screen "7161_RecipeSetpoints_STRING" 1280x715, template "7xxx_Formats"
   Button "rec_BaseScreenLocked" at 0,0 size 1280x715; TextOff 'Text'
      Visibility <- "bo_System_BaseScreenLocked"
   ScreenModuleView "Setpoint_Display_String_2" at 4,166 size 1090x44; ScreenModuleType ""
      on Guid_{11997190-50501}: function_efd93a16("pop_recipes_STRING", 200, 50, -1, -1, 1); SetTag("CPG_Recipe_Management.popupTrackers[3]", 1)
      Guid_{11997190-47977} <- "CPG_Recipe_Management.setpointsArray_STRING[1]"
      Guid_{11997190-76362} <- "[1]"
   ScreenModuleView "Setpoint_Display_String_1" at 4,132 size 1090x44; ScreenModuleType ""
      on Guid_{11997190-50501}: function_efd93a16("pop_recipes_STRING", 200, 50, -1, -1, 1); SetTag("CPG_Recipe_Management.popupTrackers[3]", 0)
      Guid_{11997190-47977} <- "CPG_Recipe_Management.setpointsArray_STRING[0]"
      Guid_{11997190-76362} <- "[0]"
   ScreenModuleView "Setpoint_Display_String_3" at 4,200 size 1090x44; ScreenModuleType ""
      on Guid_{11997190-50501}: function_efd93a16("pop_recipes_STRING", 200, 50, -1, -1, 1); SetTag("CPG_Recipe_Management.popupTrackers[3]", 2)
      Guid_{11997190-47977} <- "CPG_Recipe_Management.setpointsArray_STRING[2]"
      Guid_{11997190-76362} <- "[2]"
   ScreenModuleView "Setpoint_Display_String_4" at 4,234 size 1090x44; ScreenModuleType ""
      on Guid_{11997190-50501}: function_efd93a16("pop_recipes_STRING", 200, 50, -1, -1, 1); SetTag("CPG_Recipe_Management.popupTrackers[3]", 3)
      Guid_{11997190-47977} <- "CPG_Recipe_Management.setpointsArray_STRING[3]"
      Guid_{11997190-76362} <- "[3]"
   ScreenModuleView "Setpoint_Display_String_5" at 4,268 size 1090x44; ScreenModuleType ""
      on Guid_{11997190-50501}: function_efd93a16("pop_recipes_STRING", 200, 50, -1, -1, 1); SetTag("CPG_Recipe_Management.popupTrackers[3]", 4)
      Guid_{11997190-47977} <- "CPG_Recipe_Management.setpointsArray_STRING[4]"
      Guid_{11997190-76362} <- "[4]"
   ScreenModuleView "Setpoint_Display_String_6" at 4,302 size 1090x44; ScreenModuleType ""
      on Guid_{11997190-50501}: function_efd93a16("pop_recipes_STRING", 200, 50, -1, -1, 1); SetTag("CPG_Recipe_Management.popupTrackers[3]", 5)
      Guid_{11997190-47977} <- "CPG_Recipe_Management.setpointsArray_STRING[5]"
      Guid_{11997190-76362} <- "[5]"
   ScreenModuleView "Setpoint_Display_String_7" at 4,336 size 1090x44; ScreenModuleType ""
      on Guid_{11997190-50501}: function_efd93a16("pop_recipes_STRING", 200, 50, -1, -1, 1); SetTag("CPG_Recipe_Management.popupTrackers[3]", 6)
      Guid_{11997190-47977} <- "CPG_Recipe_Management.setpointsArray_STRING[6]"
      Guid_{11997190-76362} <- "[6]"
   ScreenModuleView "Setpoint_Display_String_8" at 4,370 size 1090x44; ScreenModuleType ""
      on Guid_{11997190-50501}: function_efd93a16("pop_recipes_STRING", 200, 50, -1, -1, 1); SetTag("CPG_Recipe_Management.popupTrackers[3]", 7)
      Guid_{11997190-47977} <- "CPG_Recipe_Management.setpointsArray_STRING[7]"
      Guid_{11997190-76362} <- "[7]"
   ScreenModuleView "Setpoint_Display_String_9" at 4,404 size 1090x44; ScreenModuleType ""
      on Guid_{11997190-50501}: function_efd93a16("pop_recipes_STRING", 200, 50, -1, -1, 1); SetTag("CPG_Recipe_Management.popupTrackers[3]", 8)
      Guid_{11997190-47977} <- "CPG_Recipe_Management.setpointsArray_STRING[8]"
      Guid_{11997190-76362} <- "[8]"
   ScreenModuleView "Setpoint_Display_String_10" at 4,438 size 1090x44; ScreenModuleType ""
      on Guid_{11997190-50501}: function_efd93a16("pop_recipes_STRING", 200, 50, -1, -1, 1); SetTag("CPG_Recipe_Management.popupTrackers[3]", 9)
      Guid_{11997190-47977} <- "CPG_Recipe_Management.setpointsArray_STRING[9]"
      Guid_{11997190-76362} <- "[9]"
   ScreenModuleView "Setpoint_Display_String_11" at 4,472 size 1090x44; ScreenModuleType ""
      on Guid_{11997190-50501}: function_efd93a16("pop_recipes_STRING", 200, 50, -1, -1, 1); SetTag("CPG_Recipe_Management.popupTrackers[3]", 10)
      Guid_{11997190-47977} <- "CPG_Recipe_Management.setpointsArray_STRING[10]"
      Guid_{11997190-76362} <- "[10]"
   ScreenModuleView "Setpoint_Display_String_12" at 4,506 size 1090x44; ScreenModuleType ""
      on Guid_{11997190-50501}: function_efd93a16("pop_recipes_STRING", 200, 50, -1, -1, 1); SetTag("CPG_Recipe_Management.popupTrackers[3]", 11)
      Guid_{11997190-47977} <- "CPG_Recipe_Management.setpointsArray_STRING[11]"
      Guid_{11997190-76362} <- "[11]"
   TextField "Text field_9" at 125,40 size 227x25; Text 'RECIPE SETPOINTS - STRING / Rezeptur Sollwerte - STRING'
   Button "Button_3" at 160,555 size 78x45; TextOff 'Text'; PictureOff "Up_Arrow"
      on Release: function_b9b71300("CPG_Recipe_Management.currentPages[3]", 1)
   Button "Button_4" at 287,555 size 78x45; TextOff 'Text'; PictureOff "Down_Arrow"
      on Release: function_dd21b452("CPG_Recipe_Management.currentPages[3]", 1)
   TextField "Text field_10" at 35,565 size 126x25; Text 'Pg Up/Down / Seite vor/zurück'
   IOField "I/O field_3" at 446,565 size 35x25; FormatPattern 999
      ProcessValue <- "CPG_Recipe_Management.currentPages[3]"
   TextField "Text field_13" at 381,565 size 60x25; Text 'Page # / Seite #'
   TextField "Text field_14" at 488,565 size 32x25; Text 'of / von'
   IOField "I/O field_4" at 534,564 size 37x27; FormatPattern 999
      ProcessValue <- "CPG_Recipe_Management.maxPages[3]"
   TextField "Text field_2" at 35,93 size 115x25; Text 'Setpoint Name / Sollwert-Name'
   TextField "Text field_6" at 243,83 size 72x46; Text 'Current Value Aktueller Wert'
   TextField "Text field_7" at 384,93 size 32x25; Text 'Min'
   TextField "Text field_4" at 506,93 size 36x25; Text 'Max'
   IOField "I/O field_9" at 757,42 size 53x36; FormatPattern 999
      ProcessValue <- "RecipeID_A"
   IOField "I/O field_10" at 883,42 size 53x36; FormatPattern 999
      ProcessValue <- "RecipeID_B"
   IOField "I/O field_11" at 998,42 size 53x36; FormatPattern 999
      ProcessValue <- "RecipeID_C"
   IOField "I/O field_13" at 550,83 size 187x22; FormatPattern ????????????????????
      ProcessValue <- "CurrentRecipeName"
   IOField "I/O field_14" at 907,104 size 187x22; FormatPattern ????????????????????
      ProcessValue <- "RecipeName_C"
   IOField "I/O field_15" at 816,83 size 187x22; FormatPattern ????????????????????
      ProcessValue <- "RecipeName_B"
   IOField "I/O field_16" at 690,103 size 187x23; FormatPattern ????????????????????
      ProcessValue <- "RecipeName_A"
   TextField "Text field_1" at 748,15 size 98x25; Text 'Recipe A / Datensatz A'
   TextField "Text field_3" at 874,15 size 97x25; Text 'Recipe B / Datensatz B'
   TextField "Text field_8" at 989,15 size 97x25; Text 'Recipe C / Datensatz C'
   Group "Group" at 588,37 size 110x46
   TextField "Text field_5" at 588,37 size 88x46; Text 'Current Recipe: Aktueller Datensatz:'
   IOField "I/O field_12" at 663,48 size 35x25; FormatPattern 999
      ProcessValue <- "CurrentRecipeID"

screen "6001_SystemDiagnostic" 1280x715, template "6xxx_Diagnostics"
   SysDiagControl "ctrlSystemDiagnostics" at 15,15 size 1035x595
   Button "btnSystemDiagnosticsVerticalScrollUp" at 1050,70 size 40x30; TextOff 'Text'; PictureOff "icn-scroll-up-20x11"
      on Release: function_b22acb07("ctrlSystemDiagnostics")
   Button "btnSystemDiagnosticsVerticalScrollDown" at 1050,529 size 40x30; TextOff 'Text'; PictureOff "icn-scroll-down-20x11"
      on Release: function_b8b2ebe3("ctrlSystemDiagnostics")
   SysDiagControl "ctrlSystemDiagnosticsLocked" at 15,15 size 1035x595
      Visibility <- "bo_System_BaseScreenLocked"
   Rectangle "recBaseScreenLocked" at 0,0 size 1280x708
      Visibility <- "bo_System_BaseScreenLocked"

screen "6041_WebDiagnostic" 1280x715, template "6xxx_Diagnostics"
   HTMLBrowser "ctrlHTMLBrowser" at 16,16 size 1073x531
      Address <- "str_Diagnostic_WebURL"
   Button "btnWebServerPLC" at 15,560 size 125x50; TextOff 'PLC / SPS'
      on Release: SetTag("str_Diagnostic_WebURL", '192.168.0.1')
   Rectangle "recBaseScreenLocked" at 0,0 size 1280x708
      Visibility <- "bo_System_BaseScreenLocked"

Template "1xxx_MachineControl" 1280x715
   ScreenModuleView "fcpBodyBar" at 5,5 size 1270x615; Guid_{11997190-53329} 'Up & Downstream'; Guid_{11997190-53335} 'OMAC Times OMAC Zeiten Timers / OEE'; Guid_{11997190-53325} 'Overview / Übersicht / Equipment view'; Guid_{11997190-53331} 'OMAC State Model OMAC Statusmodell OMAC State Model'; Guid_{11997190-53337} 'OEE / Manual CMD's'; Guid_{11997190-53333} 'OMAC PackTags PackTags'; Guid_{11997190-53339} 'Manual Commands Manuelle Kommandos PDI Interface'; ScreenModuleType ""
      on Guid_{11997190-53582}: ActivateScreen("1201_OEE", 0)
      on Guid_{11997190-53576}: ActivateScreen("1081_OMACStateModel", 0)
      on Guid_{11997190-53580}: ActivateScreen("1161_OMACTimes", 0)
      on Guid_{11997190-53584}: ActivateScreen("1241_ManualCommands", 0)
      on Guid_{11997190-53578}: ActivateScreen("1121_OMACPackTags", 0)
      on Guid_{11997190-53574}: ActivateScreen("1041_Up&Downstream", 0)
      on Guid_{11997190-53572}: ActivateScreen("1001_EquipmentView1", 0)
      Guid_{11997190-62386} <- "HMI_Data.HMICurrentScreenID"
      Guid_{11997190-53044} <- "i16_1000_MachineControl_SecondNavMaxTopics"
   ScreenModuleView "fcpBottomBar" at 5,625 size 1270x85; ScreenModuleType ""
      on Guid_{11997190-126458}: function_efd93a16("pop_UserLogin", 437, 285, 1, -1, 1)
      on Guid_{11997190-96858}: ActivateScreen("6001_SystemDiagnostic", 0)
      on Guid_{11997190-96860}: ActivateScreen("7001_RecipeControl", 0)
      on Guid_{11997190-126452}: "sub_OpenPrevScreen"()
      on Guid_{11997190-96848}: ActivateScreen("1001_EquipmentView1", 0)
      on Guid_{11997190-96850}: ActivateScreen("2001_Settings", 0)
      on Guid_{11997190-96852}: ActivateScreen("3001_AlarmOverview", 0)
      Guid_{11997190-60598} <- "HMI_Data.HMICurrentScreenID"
   Button "btnCntrlCmdStart" at 835,638 size 70x70; TextOff 'Text'; PictureOff "icn-omac-start"
      on Release: ResetBit("HMI_Data.CMDs.PB_Start")
      on Press: SetBit("HMI_Data.CMDs.PB_Start")
      Appearance <- "HMI_Data.CMDs.PB_Start"
   Button "btnCntrlCmdStop" at 910,638 size 70x70; TextOff 'Text'; PictureOff "icn-omac-stop"
      on Release: ResetBit("HMI_Data.CMDs.PB_Stop")
      on Press: SetBit("HMI_Data.CMDs.PB_Stop")
      Appearance <- "HMI_Data.CMDs.PB_Stop"
   Button "btnCntrlCmdReset" at 985,638 size 70x70; TextOff 'Text'; PictureOff "icn-omac-reset"
      on Release: ResetBit("HMI_Data.CMDs.PB_Reset")
      on Press: SetBit("HMI_Data.CMDs.PB_Reset")
      Appearance <- "HMI_Data.CMDs.PB_Reset"
   Switch "Switch_EStop" at 1126,517 size 132x58; CaptionText 'Switch'; TextOff 'E-Stop Released Not-Halt Quittiert'; TextOn 'E-Stop Pressed Not-Halt Aktiv'
      ProcessValue <- "HMI_Data_CPG.CMDs.PB_EStop"
      Appearance <- "HMI_Data_CPG.CMDs.PB_EStop"

Template "2xxx_Settings" 1280x715
   ScreenModuleView "fcpBodyBar" at 5,5 size 1270x615; Guid_{11997190-53325} 'Station A / Estacion A'; Guid_{11997190-53331} 'Benutzer- verwaltung'; Guid_{11997190-53329} 'System Functions System- funktionen Estacion B'; ScreenModuleType ""
      on Guid_{11997190-53576}: ActivateScreen("2081_UserManagement", 0)
      on Guid_{11997190-53574}: ActivateScreen("2041_SystemFunctions", 0)
      on Guid_{11997190-53572}: ActivateScreen("2001_Settings", 0)
      Guid_{11997190-62386} <- "HMI_Data.HMICurrentScreenID"
      Guid_{11997190-53044} <- "i16_2000_Settings_SecondNavMaxTopics"
   ScreenModuleView "fcpBottomBar" at 5,625 size 1270x85; ScreenModuleType ""
      on Guid_{11997190-126458}: function_efd93a16("pop_UserLogin", 437, 285, 1, -1, 1)
      on Guid_{11997190-96858}: ActivateScreen("6001_SystemDiagnostic", 0)
      on Guid_{11997190-96860}: ActivateScreen("7001_RecipeControl", 0)
      on Guid_{11997190-126452}: "sub_OpenPrevScreen"()
      on Guid_{11997190-96848}: ActivateScreen("1001_EquipmentView1", 0)
      on Guid_{11997190-96850}: ActivateScreen("2001_Settings", 0)
      on Guid_{11997190-96852}: ActivateScreen("3001_AlarmOverview", 0)
      Guid_{11997190-60598} <- "HMI_Data.HMICurrentScreenID"
   Button "btnCntrlCmdStart" at 835,638 size 70x70; TextOff 'Text'; PictureOff "icn-omac-start"
      on Release: ResetBit("HMI_Data.CMDs.PB_Start")
      on Press: SetBit("HMI_Data.CMDs.PB_Start")
      Appearance <- "HMI_Data.CMDs.PB_Start"
   Button "btnCntrlCmdStop" at 910,638 size 70x70; TextOff 'Text'; PictureOff "icn-omac-stop"
      on Release: ResetBit("HMI_Data.CMDs.PB_Stop")
      on Press: SetBit("HMI_Data.CMDs.PB_Stop")
      Appearance <- "HMI_Data.CMDs.PB_Stop"
   Button "btnCntrlCmdReset" at 985,638 size 70x70; TextOff 'Text'; PictureOff "icn-omac-reset"
      on Release: ResetBit("HMI_Data.CMDs.PB_Reset")
      on Press: SetBit("HMI_Data.CMDs.PB_Reset")
      Appearance <- "HMI_Data.CMDs.PB_Reset"

Template "3xxx_Alarms&Events" 1280x715
   ScreenModuleView "fcpBodyBar" at 5,5 size 1270x615; Guid_{11997190-53329} 'Alarm Events / Alarmmeldungen'; Guid_{11997190-53335} 'Pareto Alarm Tracking'; Guid_{11997190-53325} 'Event Overview / Meldeübersicht'; Guid_{11997190-53331} 'Warning Events / Warnmeldungen / Eventos de advertencia'; Guid_{11997190-53333} 'HMI Events / HMI Meldungen'; ScreenModuleType ""
      on Guid_{11997190-53576}: ActivateScreen("3081_WarningEvents", 0)
      on Guid_{11997190-53574}: ActivateScreen("3041_AlarmEvents", 0)
      on Guid_{11997190-53578}: ActivateScreen("3121_HMI_Alarms", 0)
      on Guid_{11997190-53580}: ActivateScreen("3161_ParetoAlarmData", 0)
      on Guid_{11997190-53572}: ActivateScreen("3001_AlarmOverview", 0)
      Guid_{11997190-62386} <- "HMI_Data.HMICurrentScreenID"
      Guid_{11997190-53044} <- "i16_3000_Alarms&Events_SecondNavMaxTopics"
   ScreenModuleView "fcpBottomBar" at 5,625 size 1270x85; ScreenModuleType ""
      on Guid_{11997190-126458}: function_efd93a16("pop_UserLogin", 437, 285, 1, -1, 1)
      on Guid_{11997190-96858}: ActivateScreen("6001_SystemDiagnostic", 0)
      on Guid_{11997190-96860}: ActivateScreen("7001_RecipeControl", 0)
      on Guid_{11997190-126452}: "sub_OpenPrevScreen"()
      on Guid_{11997190-96848}: ActivateScreen("1001_EquipmentView1", 0)
      on Guid_{11997190-96850}: ActivateScreen("2001_Settings", 0)
      on Guid_{11997190-96852}: ActivateScreen("3001_AlarmOverview", 0)
      Guid_{11997190-60598} <- "HMI_Data.HMICurrentScreenID"
   Button "btnCntrlCmdStart" at 835,638 size 70x70; TextOff 'Text'; PictureOff "icn-omac-start"
      on Release: ResetBit("HMI_Data.CMDs.PB_Start")
      on Press: SetBit("HMI_Data.CMDs.PB_Start")
      Appearance <- "HMI_Data.CMDs.PB_Start"
   Button "btnCntrlCmdStop" at 910,638 size 70x70; TextOff 'Text'; PictureOff "icn-omac-stop"
      on Release: ResetBit("HMI_Data.CMDs.PB_Stop")
      on Press: SetBit("HMI_Data.CMDs.PB_Stop")
      Appearance <- "HMI_Data.CMDs.PB_Stop"
   Button "btnCntrlCmdReset" at 985,638 size 70x70; TextOff 'Text'; PictureOff "icn-omac-reset"
      on Release: ResetBit("HMI_Data.CMDs.PB_Reset")
      on Press: SetBit("HMI_Data.CMDs.PB_Reset")
      Appearance <- "HMI_Data.CMDs.PB_Reset"

Template "6xxx_Diagnostics" 1280x715
   ScreenModuleView "fcpBodyBar" at 5,5 size 1270x615; Guid_{11997190-53325} 'System Diagnostic System- diagnose Diagnóstico del sistema'; Guid_{11997190-53329} 'Web Diagnostic Web- diagnose Diagnóstico web'; ScreenModuleType ""
      on Guid_{11997190-53574}: ActivateScreen("6041_WebDiagnostic", 0)
      on Guid_{11997190-53572}: ActivateScreen("6001_SystemDiagnostic", 0)
      Guid_{11997190-62386} <- "HMI_Data.HMICurrentScreenID"
      Guid_{11997190-53044} <- "i16_6000_Diagnostics_SecondNavMaxTopics"
   ScreenModuleView "fcpBottomBar" at 5,625 size 1270x85; ScreenModuleType ""
      on Guid_{11997190-126458}: function_efd93a16("pop_UserLogin", 437, 285, 1, -1, 1)
      on Guid_{11997190-96858}: ActivateScreen("6001_SystemDiagnostic", 0)
      on Guid_{11997190-96860}: ActivateScreen("7001_RecipeControl", 0)
      on Guid_{11997190-126452}: "sub_OpenPrevScreen"()
      on Guid_{11997190-96848}: ActivateScreen("1001_EquipmentView1", 0)
      on Guid_{11997190-96850}: ActivateScreen("2001_Settings", 0)
      on Guid_{11997190-96852}: ActivateScreen("3001_AlarmOverview", 0)
      Guid_{11997190-60598} <- "HMI_Data.HMICurrentScreenID"
   Button "btnCntrlCmdStart" at 835,638 size 70x70; TextOff 'Text'; PictureOff "icn-omac-start"
      on Release: ResetBit("HMI_Data.CMDs.PB_Start")
      on Press: SetBit("HMI_Data.CMDs.PB_Start")
      Appearance <- "HMI_Data.CMDs.PB_Start"
   Button "btnCntrlCmdStop" at 910,638 size 70x70; TextOff 'Text'; PictureOff "icn-omac-stop"
      on Release: ResetBit("HMI_Data.CMDs.PB_Stop")
      on Press: SetBit("HMI_Data.CMDs.PB_Stop")
      Appearance <- "HMI_Data.CMDs.PB_Stop"
   Button "btnCntrlCmdReset" at 985,638 size 70x70; TextOff 'Text'; PictureOff "icn-omac-reset"
      on Release: ResetBit("HMI_Data.CMDs.PB_Reset")
      on Press: SetBit("HMI_Data.CMDs.PB_Reset")
      Appearance <- "HMI_Data.CMDs.PB_Reset"

Template "7xxx_Formats" 1280x715
   ScreenModuleView "fcpBodyBar" at 5,5 size 1270x615; Guid_{11997190-53329} 'REAL Sollwerte'; Guid_{11997190-53335} 'STRING Sollwerte'; Guid_{11997190-53325} 'Recipe Control Rezepturverwaltung'; Guid_{11997190-53331} 'DINT Sollwerte'; Guid_{11997190-53333} 'BOOL Sollwerte'; ScreenModuleType ""
      on Guid_{11997190-53576}: ActivateScreen("7081_RecipeSetpoints_DINT", 0)
      on Guid_{11997190-53580}: ActivateScreen("7161_RecipeSetpoints_STRING", 0)
      on Guid_{11997190-53578}: ActivateScreen("7121_RecipeSetpoints_BOOL", 0)
      on Guid_{11997190-53574}: ActivateScreen("7041_RecipeSetpoints_REAL", 0)
      on Guid_{11997190-53572}: ActivateScreen("7001_RecipeControl", 0)
      Guid_{11997190-62386} <- "HMI_Data.HMICurrentScreenID"
      Guid_{11997190-53044} <- "i16_7000_Formats_SecondNavMaxTopics"
   ScreenModuleView "fcpBottomBar" at 5,625 size 1270x85; ScreenModuleType ""
      on Guid_{11997190-126458}: function_efd93a16("pop_UserLogin", 437, 285, 1, -1, 1)
      on Guid_{11997190-96858}: ActivateScreen("6001_SystemDiagnostic", 0)
      on Guid_{11997190-96860}: ActivateScreen("7001_RecipeControl", 0)
      on Guid_{11997190-126452}: "sub_OpenPrevScreen"()
      on Guid_{11997190-96848}: ActivateScreen("1001_EquipmentView1", 0)
      on Guid_{11997190-96850}: ActivateScreen("2001_Settings", 0)
      on Guid_{11997190-96852}: ActivateScreen("3001_AlarmOverview", 0)
      Guid_{11997190-60598} <- "HMI_Data.HMICurrentScreenID"
   Button "btnCntrlCmdStart" at 835,638 size 70x70; TextOff 'Text'; PictureOff "icn-omac-start"
      on Release: ResetBit("HMI_Data.CMDs.PB_Start")
      on Press: SetBit("HMI_Data.CMDs.PB_Start")
      Appearance <- "HMI_Data.CMDs.PB_Start"
   Button "btnCntrlCmdStop" at 910,638 size 70x70; TextOff 'Text'; PictureOff "icn-omac-stop"
      on Release: ResetBit("HMI_Data.CMDs.PB_Stop")
      on Press: SetBit("HMI_Data.CMDs.PB_Stop")
      Appearance <- "HMI_Data.CMDs.PB_Stop"
   Button "btnCntrlCmdReset" at 985,638 size 70x70; TextOff 'Text'; PictureOff "icn-omac-reset"
      on Release: ResetBit("HMI_Data.CMDs.PB_Reset")
      on Press: SetBit("HMI_Data.CMDs.PB_Reset")
      Appearance <- "HMI_Data.CMDs.PB_Reset"

PopupScreen "pop_ErrorScreenNo" 405x230
   on GenerateScreen: SetBit("bo_System_BaseScreenLocked")
   on ClearScreen: ResetBit("bo_System_BaseScreenLocked")
   Button "btnClose" at 140,170 size 125x50; TextOff 'Close / Schließen'
      on Click: function_efd93a16("pop_ErrorScreenNo", 0, 0, 0, -1, 1)
   TextField "txtMessage" at 10,65 size 390x105; Text 'The screen number could not be determined! Please check the screen name. Die Bildnummer konnte nicht ermittelt werden! Bitte überprüfen Sie den Bildnamen. The Screen name has the wrong Style'
   Button "btnHeader" at 3,3 size 399x60; TextOff 'System Error / Systemfehler'

PopupScreen "pop_UserLogin" 405x230
   on GenerateScreen: SetBit("bo_System_BaseScreenLocked")
   on ClearScreen: ResetBit("bo_System_BaseScreenLocked")
   Button "btnLogOff" at 10,170 size 125x50; TextOff 'Log off / Ausloggen / Desconectarse'
      on Release: function_efd93a16("pop_UserLogin", 0, 0, 0, -1, 1); function_f23ef4c9()
   Button "btnChangeUser" at 140,170 size 125x50; TextOff 'Change User Benutzer- wechsel'
      on Release: function_efd93a16("pop_UserLogin", 0, 0, 0, -1, 1); function_a2a04561()
   Button "btnClose" at 270,170 size 125x50; TextOff 'Close / Schließen'
      on Release: function_efd93a16("pop_UserLogin", 0, 0, 0, -1, 1)
   TextField "txtMessage" at 10,65 size 390x105; Text 'Log off or change user? / Ausloggen oder Benutzerwechsel?'
   Button "btnHeader" at 3,3 size 399x60; TextOff 'User Management / Benutzerverwaltung'

PopupScreen "pop_recipes_BOOL" 645x584
   ScreenModuleView "Bool Popup_1_1" at 2,1 size 640x579; ScreenModuleType ""
      on Guid_{11997190-50035}: ActivateScreen("7121_RecipeSetpoints_BOOL", 0)
      Guid_{11997190-48328} <- "CPG_Recipe_Management.setpointPopup_BOOL"
      Guid_{11997190-42630} <- "CPG_RecipeCfg.recipeControl"

PopupScreen "pop_recipes_DINT" 645x584
   ScreenModuleView "Dint Popup_1" at 0,0 size 640x579; ScreenModuleType ""
      on Guid_{11997190-50035}: ActivateScreen("7081_RecipeSetpoints_DINT", 0)
      Guid_{11997190-48328} <- "CPG_Recipe_Management.setpointPopup_DINT"
      Guid_{11997190-42630} <- "CPG_RecipeCfg.recipeControl"

PopupScreen "pop_recipes_REAL" 642x581
   ScreenModuleView "Real Popup_1" at 0,0 size 640x579; ScreenModuleType ""
      on Guid_{11997190-50035}: ActivateScreen("7041_RecipeSetpoints_REAL", 0)
      Guid_{11997190-48328} <- "CPG_Recipe_Management.setpointPopup_REAL"
      Guid_{11997190-42630} <- "CPG_RecipeCfg.recipeControl"

PopupScreen "pop_recipes_STRING" 645x584
   ScreenModuleView "Popup_String_1" at 2,0 size 640x579; ScreenModuleType ""
      on Guid_{11997190-50035}: ActivateScreen("7161_RecipeSetpoints_STRING", 0)
      Guid_{11997190-48328} <- "CPG_Recipe_Management.setpointPopup_STRING"
      Guid_{11997190-42630} <- "CPG_RecipeCfg.recipeControl"

VB script "sub_SetScreenBrightness"
   '****************************************************************************************************************************
   '----------------------------------------------------------------------------------------------------------------------------
   ' Functionality : Changing the screen brightness with a defined increment size
   ' Run           : After a user change via the task scheduler
   ' Run system    : WinCC Comfort/Advanced Runtime V13
   '----------------------------------------------------------------------------------------------------------------------------
   ' Script parameters:
   '  Parameter        | Data type    | Description
   '  i16Offset        | INTEGER      | Specifies the increment by which the screen brightness is changed
   '----------------------------------------------------------------------------------------------------------------------------
   ' Change table:
   '  Version    | Date     | Creator         | Description
   '  01.00.00   | 18/06/18 | Briese, Mike    | Creation
   '----------------------------------------------------------------------------------------------------------------------------
   '****************************************************************************************************************************
   
   'Declaration
   Dim i16NewDisplayBrightness
   
   
   'Determine new value for screen brightness
   i16NewDisplayBrightness = SmartTags("i16_Settings_CurDisplayBrightness") + i16Offset
   
   'Check whether new value is within the limits
   '=> If No, then set to the corresponding limit value
   If i16NewDisplayBrightness < 20 Then
   	i16NewDisplayBrightness = 20
   ElseIf i16NewDisplayBrightness > 100 Then
   	i16NewDisplayBrightness = 100
   End If
   
   'Take over new value
   SmartTags("i16_Settings_CurDisplayBrightness") = i16NewDisplayBrightness
   e4c2bb66-d114-4215-9f74-4e7e992fb119 i16NewDisplayBrightness

VB script "sub_ScreenChanged"
   '****************************************************************************************************************************
   '----------------------------------------------------------------------------------------------------------------------------
   ' Functionality : Determining the screen number from the screen name
   ' Run           : After a screen change via the task scheduler
   ' Run system    : WinCC Comfort/Advanced Runtime V13
   '----------------------------------------------------------------------------------------------------------------------------
   ' Script parameters:
   '  Parameter        | Data type    | Description
   '                   |              |
   '----------------------------------------------------------------------------------------------------------------------------
   ' Change table:
   '  Version    | Date     | Creator         | Description
   '  01.00.00   | 18/06/18 | Briese, Mike    | Creation
   '----------------------------------------------------------------------------------------------------------------------------
   '****************************************************************************************************************************
   
   'Declaration
   Dim strCurScreenName, i16NewScreenID, i16Index
   
   
   'Determine screen number from screen name
   strCurScreenName = HmiRuntime.BaseScreenName
   i16NewScreenID = Mid(strCurScreenName, 1, 4)
   
   'Plausibility check of the determined screen number
   '=> if it is not plausible, show an error message and exit sub
   If Not IsNumeric(i16NewScreenID) Then
   	efd93a16-2665-4b85-bcb9-25eddcb7b6f4 pop_ErrorScreenNo, 437, 285, $3$hmiOn$, $3$hmiAnimationOff$, $3$hmiMedium$
   	SmartTags("HMI_Data.HMICurrentScreenID") = -1
   	Exit Sub
   End If 
   
   'Take over determined screen number
   SmartTags("HMI_Data.HMICurrentScreenID") = i16NewScreenID
   
   'Take over determined screen number to screen buffer for return function, if this is not active
   i16Index = SmartTags("i16_System_PrevScreenPointer")
   If SmartTags("bo_System_PrevScreenActive") Then
   	SmartTags("bo_System_PrevScreenActive") = False
   Else
   	If i16Index < UBound(SmartTags("arr_System_PrevScreenStorage")) Then
   		i16Index = i16Index + 1
   	Else
   		i16Index = 0
   	End If
   	SmartTags("i16_System_PrevScreenPointer") = i16Index
   	SmartTags("arr_System_PrevScreenStorage")(i16Index) = i16NewScreenID
   End If

VB script "sub_RuntimeStart"
   '****************************************************************************************************************************
   '----------------------------------------------------------------------------------------------------------------------------
   ' Functionality : This script contains all one-time actions that are to be executed after the runtime start
   ' Run           : Runtime start of HMI project
   ' Run system    : WinCC Comfort/Advanced Runtime V13
   '----------------------------------------------------------------------------------------------------------------------------
   ' Script parameters:
   '  Parameter        | Data type    | Description
   '                   |              |
   '----------------------------------------------------------------------------------------------------------------------------
   ' Change table:
   '  Version    | Date     | Creator         | Description
   '  01.00.00   | 18/06/18 | Briese, Mike    | Creation
   '----------------------------------------------------------------------------------------------------------------------------
   '****************************************************************************************************************************
   
   
   'Determine current user info
   sub_UserChanged
   
   'Open overview screen
   bec8f1e5-2ab1-45f6-ad91-1d37c469eb91 1001_EquipmentView1, 0

VB script "sub_OpenPrevScreen"
   '****************************************************************************************************************************
   '----------------------------------------------------------------------------------------------------------------------------
   ' Functionality : Open previous screen
   '                 An screen buffer is required for this function. 
   ' Run           : On demand
   ' Run system    : WinCC Comfort/Advanced Runtime V13
   '----------------------------------------------------------------------------------------------------------------------------
   ' Script parameters:
   '  Parameter        | Data type    | Description
   '                   |              |
   '----------------------------------------------------------------------------------------------------------------------------
   ' Change table:
   '  Version    | Date     | Creator         | Description
   '  01.00.00   | 18/06/18 | Briese, Mike    | Creation
   '----------------------------------------------------------------------------------------------------------------------------
   '****************************************************************************************************************************
   
   'Declaration
   Const strFctName = "sub_OpenPrevScreen"
   Dim i16CurBufferIndex, i16NewBufferIndex, i16ScreenID
   
   
   'Load number of previous screen from screen buffer
   i16CurBufferIndex = SmartTags("i16_System_PrevScreenPointer")
   If i16CurBufferIndex > 0 Then
   	i16NewBufferIndex = i16CurBufferIndex - 1
   Else
   	i16NewBufferIndex = UBound(SmartTags("arr_System_PrevScreenStorage"))
   End If
   
   'Check if screen buffer element contains a valid number
   '=> if no, then the function is terminated
   i16ScreenID = SmartTags("arr_System_PrevScreenStorage")(i16NewBufferIndex)
   If i16ScreenID = 0 Then Exit Sub
   
   'Reset current screen buffer element and accept new pointer
   SmartTags("arr_System_PrevScreenStorage")(i16CurBufferIndex) = 0
   SmartTags("i16_System_PrevScreenPointer") = i16NewBufferIndex
   
   'Set auxiliary flag for screen change function
   SmartTags("bo_System_PrevScreenActive") = True
   
   'Open previous screen
   acd163fa-ee86-4170-88da-c8d9ec58660c i16ScreenID, 0

VB script "sub_UserChanged"
   '****************************************************************************************************************************
   '----------------------------------------------------------------------------------------------------------------------------
   ' Functionality : Determining the screen number from the screen name
   '                 The associated group number/name and authorizations are determined according to the current user selection.
   '                 Afterwards, a '0' is entered at the current pointer position in the screen storage for the return function,
   '                 so that the new user cannot jump to the last called screens of the previous user. Finally, the overview
   '                 screen is opened.
   ' Run           : After a user change via the task scheduler
   ' Run system    : WinCC Comfort/Advanced Runtime V13
   '----------------------------------------------------------------------------------------------------------------------------
   ' Script parameters:
   '  Parameter        | Data type    | Description
   '                   |              |
   '----------------------------------------------------------------------------------------------------------------------------
   ' Change table:
   '  Version    | Date     | Creator         | Description
   '  01.00.00   | 18/06/18 | Briese, Mike    | Creation
   '----------------------------------------------------------------------------------------------------------------------------
   '****************************************************************************************************************************
   
   'Declaration
   Dim arrUserName, strUserName(2), strUserNamePart1, strUserNamePart2, strLoginData
   Dim i16Index
   
   'Determine current user name
   f41c6f6c-971d-4734-9362-16d81ac70597 str_System_CurUser
   If SmartTags("str_System_CurUser") = "" Then
   	SmartTags("str_System_CurUser") = "-"
   End If
   
   'Initialize current pointer index of the screen buffer for return function
   '=> to restart from here after changing users
   i16Index = SmartTags("i16_System_PrevScreenPointer")
   SmartTags("arr_System_PrevScreenStorage")(i16Index) = 0
   
   'Reset basic screen lock
   '=> required if incorrect login data has been entered
   SmartTags("bo_System_BaseScreenLocked") = False
   
   'Open overview screen
   bec8f1e5-2ab1-45f6-ad91-1d37c469eb91 1001_EquipmentView1, 0

scheduled task "ScreenChanged"
   on Action: "sub_ScreenChanged"()

scheduled task "UserChanged"
   on Action: "sub_UserChanged"()
*)

(* ===== HMI "HMI_RT_1" =====
system functions are stored by id; their names below are inferred from use

HMI tags "Default tag table"
   "testtag" : WString[10], internal

ScreenModuleEditorView "Popup_Real" 700x600
   Rectangle "Rectangle_2" at 113,186 size 434x39
      Visibility <- "Setpoint.SetpointChangeDisabled"
   TextField "NotAllowed Warning" at 131,194 size 398x23; Text 'Setpoint Changes Not Allowed in Current Machine State / Änderung im aktuellen Maschinenzustand nicht möglich'
      Visibility <- "Setpoint.SetpointChangeDisabled"
   Rectangle "Yellow" at 113,72 size 434x39
      Visibility <- "Setpoint.RecipeSetpointDiff"
   TextField "DetectDiff Warning" at 141,80 size 402x23; Text 'Current Setpoint Does Not Match Saved Recipe Value / Der aktuelle Sollwert entspricht nicht dem gespeicherten'
      Visibility <- "Setpoint.RecipeSetpointDiff"
   IOField "Current Num" at 69,346 size 46x26; FormatPattern 999
      ProcessValue <- "Control.CurrentRecipeID"
   IOField "NumA" at 69,388 size 46x26; FormatPattern 999
      ProcessValue <- "Control.RecipeID_A"
   IOField "NumB" at 69,429 size 46x26; FormatPattern 999
      ProcessValue <- "Control.RecipeID_B"
   IOField "NumC" at 69,471 size 46x26; FormatPattern 999
      ProcessValue <- "Control.RecipeID_C"
   TextField "Text field_5" at 239,305 size 112x23; Text 'Recipe Name / Datensatzname'
   TextField "Text field_6" at 517,305 size 44x23; Text 'Value / Wert'
   TextField "Text field_7" at 266,264 size 129x28; Text 'Recipe Values / Rezepturwert'
   IOField "CurrentValue_true" at 486,348 size 106x23; FormatPattern 9999999.999
      ProcessValue <- "Setpoint.CurrentRecipeValue"
   IOField "ValueA" at 486,390 size 106x25; FormatPattern 9999999.999
      ProcessValue <- "Setpoint.RecipeValueA"
   IOField "ValueB" at 486,431 size 106x23; FormatPattern 9999999.999
      ProcessValue <- "Setpoint.RecipeValueB"
   IOField "ValueC" at 486,473 size 106x23; FormatPattern 9999999.999
      ProcessValue <- "Setpoint.RecipeValueC"
   IOField "CurrentName" at 158,346 size 282x26; FormatPattern ??????????????????????????????
      ProcessValue <- "Control.CurrentRecipeName"
   IOField "NameA" at 158,388 size 282x26; FormatPattern ??????????????????????????????
      ProcessValue <- "Control.RecipeName_A"
   IOField "NameB" at 158,429 size 282x26; FormatPattern ??????????????????????????????
      ProcessValue <- "Control.RecipeName_B"
   IOField "NameC" at 158,471 size 282x26; FormatPattern ??????????????????????????????
      ProcessValue <- "Control.RecipeName_C"
   Group "Group" at 113,186 size 434x39
   Group "Group_1" at 113,72 size 434x39
   IOField "Setpoint Name" at 145,27 size 370x41; FormatPattern ????????????????????????????????
      ProcessValue <- "Setpoint.CurrentName"
   Button "Save Setpoint" at 429,233 size 154x60; TextOff 'Save Setpoint Value Sollwert Speichern'
      on Press: function_b14e0dd5("Setpoint.SaveSetpoint", 0)
   Button "Revert Setpoint" at 69,233 size 154x60; TextOff 'Revert Setpoint Value Sollwert Rücksetzen'
      on Press: function_b14e0dd5("Setpoint.RevertSetpoint", 0)
   Button "Close Button" at 79,519 size 502x60; TextOff 'CLOSE / Schließen'
   IOField "CurrentValue_true_1" at 206,153 size 132x26; FormatPattern 9999999.999
      ProcessValue <- "Setpoint.IN"
   TextField "Text field_1" at 79,307 size 36x23; Text '#'
   IOField "Max Value" at 464,154 size 106x23; FormatPattern 9999999.999
      ProcessValue <- "Setpoint.maxLimit"
   IOField "Min Value" at 93,154 size 106x23; FormatPattern 9999999.999
      ProcessValue <- "Setpoint.minLimit"
   Rectangle "Min Warning" at 94,147 size 104x36
      Visibility <- "Setpoint.minLimitReached"
   Rectangle "Max Warning" at 465,147 size 104x36
      Visibility <- "Setpoint.maxLimitReached"
   TextField "Text field_2" at 267,116 size 133x28; Text 'Current Value / Aktueller Wert'
   TextField "Text field_3" at 123,116 size 45x28; Text 'Min'
   TextField "Text field_4" at 494,116 size 45x28; Text 'Max'
   Group "Group_2" at 32,230 size 597x289
   Group "Group_3" at 345,153 size 112x23
   Rectangle "Rectangle_3" at 32,230 size 597x289
      Visibility <- "Setpoint.DisableRecipeControl"
   TextField "Text field_8" at 246,348 size 223x23; Text 'Recipe Control Disabled / Rezepturverwaltung deaktiviert'
      Visibility <- "Setpoint.DisableRecipeControl"
   TextField "Text field_10" at 345,153 size 112x23; Text '[ ]'
   IOField "Unit" at 353,153 size 96x23; FormatPattern ??????????
      ProcessValue <- "Setpoint.unit"
*)

(* ===== HMI "HMI_RT_1" =====
system functions are stored by id; their names below are inferred from use

HMI tags "Default tag table"
   "testtag" : WString[10], internal

ScreenModuleEditorView "Popup_String" 700x600
   Rectangle "Rectangle_2" at 113,154 size 434x39
      Visibility <- "Setpoint.SetpointChangeDisabled"
   TextField "NotAllowed Warning" at 131,162 size 398x23; Text 'Setpoint Changes Not Allowed in Current Machine State / Änderung im aktuellen Maschinenzustand nicht möglich'
      Visibility <- "Setpoint.SetpointChangeDisabled"
   Rectangle "Yellow" at 113,72 size 434x39
      Visibility <- "Setpoint.RecipeSetpointDiff"
   TextField "DetectDiff Warning" at 141,80 size 379x23; Text 'Current Setpoint Does Not Match Saved Recipe Value / Der aktuelle Sollwert entspricht dem gespeicherten'
      Visibility <- "Setpoint.RecipeSetpointDiff"
   IOField "Current Num" at 69,346 size 46x26; FormatPattern 999
      ProcessValue <- "Control.CurrentRecipeID"
   IOField "NumA" at 69,388 size 46x26; FormatPattern 999
      ProcessValue <- "Control.RecipeID_A"
   IOField "NumB" at 69,429 size 46x26; FormatPattern 999
      ProcessValue <- "Control.RecipeID_B"
   IOField "NumC" at 69,471 size 46x26; FormatPattern 999
      ProcessValue <- "Control.RecipeID_C"
   TextField "Text field_5" at 239,305 size 112x23; Text 'Recipe Name / Datensatzname'
   TextField "Text field_6" at 478,305 size 44x23; Text 'Value / Wert'
   TextField "Text field_7" at 266,264 size 129x28; Text 'Recipe Values / Rezepturwert'
   IOField "CurrentValue" at 453,348 size 190x23; FormatPattern ????????????????????
      ProcessValue <- "Setpoint.CurrentRecipeValue"
   IOField "ValueA" at 453,390 size 190x23; FormatPattern ????????????????????
      ProcessValue <- "Setpoint.RecipeValueA"
   IOField "ValueB" at 453,431 size 190x23; FormatPattern ????????????????????
      ProcessValue <- "Setpoint.RecipeValueB"
   IOField "ValueC" at 453,473 size 190x23; FormatPattern ????????????????????
      ProcessValue <- "Setpoint.RecipeValueC"
   IOField "CurrentName" at 158,346 size 282x26; FormatPattern ??????????????????????????????
      ProcessValue <- "Control.CurrentRecipeName"
   IOField "NameA" at 158,388 size 282x26; FormatPattern ??????????????????????????????
      ProcessValue <- "Control.RecipeName_A"
   IOField "NameB" at 158,429 size 282x26; FormatPattern ??????????????????????????????
      ProcessValue <- "Control.RecipeName_B"
   IOField "NameC" at 158,471 size 282x26; FormatPattern ??????????????????????????????
      ProcessValue <- "Control.RecipeName_C"
   Group "Group" at 113,154 size 434x39
   TextField "Text field_4" at 136,120 size 112x23; Text 'Current Value: / Aktueller Wert:'
   Group "Group_1" at 113,72 size 434x39
   IOField "Setpoint Name" at 145,27 size 370x41; FormatPattern ????????????????????????????????
      ProcessValue <- "Setpoint.CurrentSetpointName"
   Button "Save Setpoint" at 429,213 size 154x60; TextOff 'Save Setpoint Value Sollwert Speichern'
      on Press: function_b14e0dd5("Setpoint.SaveSetpoint", 0)
   Button "Revert Setpoint" at 69,213 size 154x60; TextOff 'Revert Setpoint Value Sollwert Zurücksetzen'
      on Press: function_b14e0dd5("Setpoint.RevertSetpoint", 0)
   Button "Close Button" at 79,519 size 502x60; TextOff 'CLOSE / Schließen'
   IOField "Input" at 325,119 size 192x26; FormatPattern ????????????????????
      ProcessValue <- "Setpoint.IN"
   TextField "Text field_1" at 79,307 size 36x23; Text '#'
   Group "Group_2" at 19,195 size 623x320
   Rectangle "Rectangle_3" at 19,195 size 623x320
      Visibility <- "Setpoint.DisableRecipeControl"
   TextField "Text field_2" at 242,344 size 223x23; Text 'Recipe Control Disabled / Rezepturverwaltung deaktiviert'
      Visibility <- "Setpoint.DisableRecipeControl"
*)

(* ===== HMI "HMI_RT_1" =====
system functions are stored by id; their names below are inferred from use

HMI tags "Default tag table"
   "testtag" : WString[10], internal

ScreenModuleEditorView "Popup_Dint" 700x600
   Rectangle "Yellow" at 113,72 size 434x39
      Visibility <- "Setpoint.RecipeSetpointDiff"
   TextField "DetectDiff Warning" at 141,80 size 402x23; Text 'Current Setpoint Does Not Match Saved Recipe Value / Der aktuelle Sollwert entspricht nicht dem gespeicherten'
      Visibility <- "Setpoint.RecipeSetpointDiff"
   IOField "Current Num" at 69,346 size 46x26; FormatPattern 999
      ProcessValue <- "Control.CurrentRecipeID"
   IOField "NumA" at 69,388 size 46x26; FormatPattern 999
      ProcessValue <- "Control.RecipeID_A"
   IOField "NumB" at 69,429 size 46x26; FormatPattern 999
      ProcessValue <- "Control.RecipeID_B"
   IOField "NumC" at 69,471 size 46x26; FormatPattern 999
      ProcessValue <- "Control.RecipeID_C"
   TextField "Text field_5" at 239,305 size 112x23; Text 'Recipe Name / Datensatzname'
   TextField "Text field_6" at 517,305 size 44x23; Text 'Value / Wert'
   TextField "Text field_7" at 266,264 size 129x28; Text 'Recipe Values / Rezepturwert'
   IOField "CurrentValue_true" at 491,348 size 96x23; FormatPattern 9999999999
      ProcessValue <- "Setpoint.CurrentRecipeValue"
   IOField "ValueA" at 491,390 size 96x25; FormatPattern 9999999999
      ProcessValue <- "Setpoint.RecipeValueA"
   IOField "ValueB" at 491,431 size 96x23; FormatPattern 9999999999
      ProcessValue <- "Setpoint.RecipeValueB"
   IOField "ValueC" at 491,473 size 96x23; FormatPattern 9999999999
      ProcessValue <- "Setpoint.RecipeValueC"
   IOField "CurrentName" at 158,346 size 282x26; FormatPattern ??????????????????????????????
      ProcessValue <- "Control.CurrentRecipeName"
   IOField "NameA" at 158,388 size 282x26; FormatPattern ??????????????????????????????
      ProcessValue <- "Control.RecipeName_A"
   IOField "NameB" at 158,429 size 282x26; FormatPattern ??????????????????????????????
      ProcessValue <- "Control.RecipeName_B"
   IOField "NameC" at 158,471 size 282x26; FormatPattern ??????????????????????????????
      ProcessValue <- "Control.RecipeName_C"
   Group "Group_1" at 113,72 size 434x39
   IOField "Setpoint Name" at 145,27 size 370x41; FormatPattern ????????????????????????????????
      ProcessValue <- "Setpoint.CurrentName"
   Button "Save Setpoint" at 429,233 size 154x60; TextOff 'Save Setpoint Value Sollwert Speichern'
      on Press: function_b14e0dd5("Setpoint.SaveSetpoint", 0)
   Button "Revert Setpoint" at 69,233 size 154x60; TextOff 'Revert Setpoint Value Sollwert Rücksetzen'
      on Press: function_b14e0dd5("Setpoint.RevertSetpoint", 0)
   Button "Close Button" at 79,519 size 502x60; TextOff 'CLOSE / Schließen'
   IOField "CurrentValue_true_1" at 204,153 size 132x26; FormatPattern 9999999999
      ProcessValue <- "Setpoint.IN"
   TextField "Text field_1" at 79,307 size 36x23; Text '#'
   IOField "Max Value" at 468,154 size 97x23; FormatPattern 9999999999
      ProcessValue <- "Setpoint.maxLimit"
   IOField "Min Value" at 97,154 size 97x23; FormatPattern 9999999999
      ProcessValue <- "Setpoint.minLimit"
   Rectangle "Min Warning" at 98,148 size 97x36
      Visibility <- "Setpoint.minLimitReached"
   Rectangle "Max Warning" at 469,148 size 97x36
      Visibility <- "Setpoint.maxLimitReached"
   TextField "Text field_2" at 267,116 size 133x28; Text 'Current Value / Aktueller Wert'
   TextField "Text field_3" at 123,116 size 45x28; Text 'Min'
   TextField "Text field_4" at 494,116 size 45x28; Text 'Max'
   Group "Group_2" at 26,230 size 608x289
   Group "Group" at 113,186 size 434x39
   Group "Group_3" at 346,154 size 112x23
   Rectangle "Rectangle_3" at 26,230 size 608x289
      Visibility <- "Setpoint.DisableRecipeControl"
   TextField "Text field_8" at 244,348 size 223x23; Text 'Recipe Control Disabled / Rezepturverwaltung deaktiviert'
      Visibility <- "Setpoint.DisableRecipeControl"
   Rectangle "Rectangle_2" at 113,186 size 434x39
      Visibility <- "Setpoint.SetpointChangeDisabled"
   TextField "NotAllowed Warning" at 131,194 size 398x23; Text 'Setpoint Changes Not Allowed in Current Machine State / Änderung im aktuellen Maschinenzustand nicht möglich'
      Visibility <- "Setpoint.SetpointChangeDisabled"
   IOField "Unit" at 352,154 size 100x23; FormatPattern ??????????
      ProcessValue <- "Setpoint.unit"
   TextField "Text field_10" at 346,154 size 112x23; Text '[ ]'
*)

(* ===== HMI "HMI_RT_1" =====
system functions are stored by id; their names below are inferred from use

HMI tags "Default tag table"
   "testtag" : WString[10], internal

ScreenModuleEditorView "Popup_Bool" 700x600
   Rectangle "Rectangle_2" at 113,154 size 434x39
      Visibility <- "Setpoint.SetpointChangeDisabled"
   TextField "NotAllowed Warning" at 131,162 size 398x23; Text 'Setpoint Changes Not Allowed in Current Machine State / Änderung im aktuellen Maschinenzustand nicht möglich'
      Visibility <- "Setpoint.SetpointChangeDisabled"
   Rectangle "Yellow" at 113,72 size 434x39
      Visibility <- "Setpoint.RecipeSetpointDiff"
   TextField "DetectDiff Warning" at 141,80 size 402x23; Text 'Current Setpoint Does Not Match Saved Recipe Value / Der aktuelle Sollwert entspricht nicht dem gespeicherten'
      Visibility <- "Setpoint.RecipeSetpointDiff"
   IOField "Current Num" at 69,346 size 46x26; FormatPattern 999
      ProcessValue <- "Control.CurrentRecipeID"
   IOField "NumA" at 69,388 size 46x26; FormatPattern 999
      ProcessValue <- "Control.RecipeID_A"
   IOField "NumB" at 69,429 size 46x26; FormatPattern 999
      ProcessValue <- "Control.RecipeID_B"
   IOField "NumC" at 69,471 size 46x26; FormatPattern 999
      ProcessValue <- "Control.RecipeID_C"
   TextField "Text field_5" at 239,305 size 112x23; Text 'Recipe Name / Datensatzname'
   TextField "Text field_6" at 478,305 size 44x23; Text 'Value / Wert'
   TextField "Text field_7" at 266,264 size 129x28; Text 'Recipe Values / Rezepturwert'
   IOField "CurrentValue_true" at 477,348 size 132x26; FormatPattern ??????????????
      ProcessValue <- "Setpoint.CurrentRecipeValue_Text"
   IOField "ValueA" at 474,390 size 139x26; FormatPattern ??????????????
      ProcessValue <- "Setpoint.RecipeA_Text"
   IOField "ValueB" at 478,431 size 131x26; FormatPattern ??????????????
      ProcessValue <- "Setpoint.RecipeB_Text"
   IOField "ValueC" at 478,473 size 131x26; FormatPattern ??????????????
      ProcessValue <- "Setpoint.RecipeC_Text"
   IOField "CurrentName" at 158,346 size 282x26; FormatPattern ??????????????????????????????
      ProcessValue <- "Control.CurrentRecipeName"
   IOField "NameA" at 158,388 size 282x26; FormatPattern ??????????????????????????????
      ProcessValue <- "Control.RecipeName_A"
   IOField "NameB" at 158,429 size 282x26; FormatPattern ??????????????????????????????
      ProcessValue <- "Control.RecipeName_B"
   IOField "NameC" at 158,471 size 282x26; FormatPattern ??????????????????????????????
      ProcessValue <- "Control.RecipeName_C"
   Group "Group" at 113,154 size 434x39
   TextField "Text field_4" at 134,120 size 112x23; Text 'Current Value: / Aktueller Wert:'
   Group "Group_1" at 113,72 size 434x39
   IOField "Setpoint Name" at 145,27 size 370x41; FormatPattern ????????????????????????????????
      ProcessValue <- "Setpoint.CurrentName"
   Button "Save Setpoint" at 429,213 size 154x60; TextOff 'Save Setpoint Value Sollwert Speichern'
      on Press: function_b14e0dd5("Setpoint.SaveSetpoint", 0)
   Button "Revert Setpoint" at 69,213 size 154x60; TextOff 'Revert Setpoint Value Sollwert Rücksetzen'
      on Press: function_b14e0dd5("Setpoint.RevertSetpoint", 0)
   Button "Close Button" at 79,519 size 502x60; TextOff 'CLOSE / Schließen'
   IOField "CurrentValue_true_1" at 414,120 size 152x26; FormatPattern ???????????????
      ProcessValue <- "Setpoint.Out_Text"
   Switch "Switch_1" at 267,116 size 126x33; TextOn '1'; CaptionText 'Schalter'; TextOff '0'
      ProcessValue <- "Setpoint.IN"
   TextField "Text field_1" at 79,307 size 36x23; Text '#'
   Group "Group_2" at 26,200 size 608x316
   Rectangle "Rectangle_3" at 26,200 size 608x316
      Visibility <- "Setpoint.DisableRecipeControl"
   TextField "Text field_8" at 244,344 size 219x23; Text 'Recipe Control Disabled / Rezepturverwaltung deaktviert'
      Visibility <- "Setpoint.DisableRecipeControl"
*)

(* ===== HMI "HMI_RT_1" =====

ScreenModuleEditorView "Setpoint_Display_Bool" 1200x300
   IOField "Current Recipe Value" at 603,23 size 97x23; FormatPattern ??????????
      ProcessValue <- "Data_Connection.CurrentRecipeValue_Text"
   IOField "Recipe B Value" at 855,23 size 97x23; FormatPattern ??????????
      ProcessValue <- "Data_Connection.RecipeB_Text"
   IOField "I/O field_9" at 11,15 size 190x39; FormatPattern ????????????????????
      ProcessValue <- "Data_Connection.CurrentName"
   Rectangle "Rectangle_2" at 213,23 size 121x24
      Visibility <- "Data_Connection.RecipeSetpointDiff"
   IOField "Recipe A Value" at 729,23 size 97x23; FormatPattern ??????????
      ProcessValue <- "Data_Connection.RecipeA_Text"
   IOField "Recipe C Value" at 981,23 size 97x23; FormatPattern ??????????
      ProcessValue <- "Data_Connection.RecipeC_Text"
   IOField "Current Value" at 225,23 size 97x23; FormatPattern ??????????
      ProcessValue <- "Data_Connection.Out_Text"
   TextField "Text field_1" at 380,24 size 38x22; Text 'N/A'
   TextField "Text field_2" at 506,24 size 38x22; Text 'N/A'
   Group "Group" at 338,21 size 754x28
   Button "Open Popup" at 2,21 size 1090x28; TextOff 'Text'
   Group "Group_1" at 2,21 size 1090x28
   Rectangle "Rectangle_8" at 2,21 size 1090x28
      Visibility <- "DISABLED"
   TextField "Text field_4" at 475,24 size 188x23; Text 'No Recipe Available / Kein Datensatz vorhanden'
      Visibility <- "DISABLED"
   Rectangle "Rectangle_7" at 338,21 size 754x28
      Visibility <- "Data_Connection.DisableRecipeControl"
   TextField "Text field_3" at 629,24 size 223x23; Text 'Recipe Control Disabled / Rezepturverwaltung deaktiviert'
      Visibility <- "Data_Connection.DisableRecipeControl"
*)

(* ===== HMI "HMI_RT_1" =====

ScreenModuleEditorView "Setpoint_Display_Dint" 1200x300
   IOField "Current Recipe Value" at 602,23 size 98x23; FormatPattern 9999999999
      ProcessValue <- "Data_Connection.CurrentRecipeValue"
   IOField "Recipe B Value" at 854,23 size 98x23; FormatPattern 9999999999
      ProcessValue <- "Data_Connection.RecipeValueB"
   IOField "Setpoint Name" at 11,15 size 190x39; FormatPattern ????????????????????
      ProcessValue <- "Data_Connection.CurrentName"
   Rectangle "Rectangle_2" at 211,22 size 121x24
      Visibility <- "Data_Connection.RecipeSetpointDiff"
   IOField "Recipe A Value" at 728,23 size 98x23; FormatPattern 9999999999
      ProcessValue <- "Data_Connection.RecipeValueA"
   IOField "Recipe C Value" at 980,23 size 98x23; FormatPattern 9999999999
      ProcessValue <- "Data_Connection.RecipeValueC"
   IOField "Current Value" at 224,23 size 98x23; FormatPattern 9999999999
      ProcessValue <- "Data_Connection.OUT"
   IOField "Min Value" at 350,23 size 98x23; FormatPattern 9999999999
      ProcessValue <- "Data_Connection.minLimit"
   IOField "Max Value" at 476,23 size 98x23; FormatPattern 9999999999
      ProcessValue <- "Data_Connection.maxLimit"
   Group "Group" at 338,20 size 754x28
   Button "Open Popup" at 2,20 size 1090x28; TextOff 'Text'
   Group "Group_1" at 2,20 size 1090x28
   Rectangle "Rectangle_3" at 338,20 size 754x28
      Visibility <- "Data_Connection.DisableRecipeControl"
   TextField "Text field_3" at 613,23 size 223x23; Text 'Recipe Control Disabled / Rezepturverwaltung deaktiviert'
      Visibility <- "Data_Connection.DisableRecipeControl"
   Rectangle "Rectangle_8" at 2,20 size 1090x28
      Visibility <- "DISABLED"
   TextField "Text field_1" at 475,23 size 188x23; Text 'No Recipe Available / Kein Datensatz vorhanden'
      Visibility <- "DISABLED"
*)

(* ===== HMI "HMI_RT_1" =====

ScreenModuleEditorView "Setpoint_Display_Real" 1200x300
   IOField "Current Recipe Value" at 601,23 size 100x23; FormatPattern 9999999.999
      ProcessValue <- "Data_Connection.CurrentRecipeValue"
   IOField "Recipe B Value" at 853,23 size 100x23; FormatPattern 9999999.999
      ProcessValue <- "Data_Connection.RecipeValueB"
   IOField "Setpoint Name" at 11,15 size 190x39; FormatPattern ????????????????????
      ProcessValue <- "Data_Connection.CurrentName"
   Rectangle "Rectangle_2" at 213,22 size 121x24
      Visibility <- "Data_Connection.RecipeSetpointDiff"
   IOField "Recipe A Value" at 727,23 size 100x23; FormatPattern 9999999.999
      ProcessValue <- "Data_Connection.RecipeValueA"
   IOField "Recipe C Value" at 979,23 size 100x23; FormatPattern 9999999.999
      ProcessValue <- "Data_Connection.RecipeValueC"
   IOField "Current Value" at 223,23 size 100x23; FormatPattern 9999999.999
      ProcessValue <- "Data_Connection.OUT"
   IOField "Min Value" at 349,23 size 100x23; FormatPattern 9999999.999
      ProcessValue <- "Data_Connection.minLimit"
   IOField "Max Value" at 475,23 size 100x23; FormatPattern 9999999.999
      ProcessValue <- "Data_Connection.maxLimit"
   Group "Group" at 338,20 size 754x28
   Button "Open Popup" at 2,20 size 1090x28; TextOff 'Text'
   Group "Group_1" at 2,20 size 1090x28
   Rectangle "Rectangle_3" at 338,20 size 754x28
      Visibility <- "Data_Connection.DisableRecipeControl"
   TextField "Text field_3" at 629,23 size 223x23; Text 'Recipe Control Disabled / Rezepturverwaltung deaktiviert'
      Visibility <- "Data_Connection.DisableRecipeControl"
   Rectangle "Rectangle_8" at 2,20 size 1090x28
      Visibility <- "DISABLED"
   TextField "Text field_1" at 475,23 size 188x23; Text 'No Recipe Available / Kein Datensatz vorhanden'
      Visibility <- "DISABLED"
*)

(* ===== HMI "HMI_RT_1" =====

ScreenModuleEditorView "Setpoint_Display_String" 1200x300
   IOField "Current Recipe Value" at 595,26 size 112x16; FormatPattern ????????????????????
      ProcessValue <- "Data_Connection.CurrentRecipeValue"
   IOField "Recipe B Value" at 847,26 size 112x16; FormatPattern ????????????????????
      ProcessValue <- "Data_Connection.RecipeValueB"
   IOField "I/O field_9" at 11,15 size 190x39; FormatPattern ????????????????????
      ProcessValue <- "Data_Connection.CurrentSetpointName"
   Rectangle "Rectangle_2" at 213,22 size 121x24
      Visibility <- "Data_Connection.RecipeSetpointDiff"
   IOField "Recipe A Value" at 721,26 size 112x16; FormatPattern ????????????????????
      ProcessValue <- "Data_Connection.RecipeValueA"
   IOField "Recipe C Value" at 973,26 size 112x16; FormatPattern ????????????????????
      ProcessValue <- "Data_Connection.RecipeValueC"
   IOField "Current Value" at 217,26 size 112x16; FormatPattern ????????????????????
      ProcessValue <- "Data_Connection.OUT"
   TextField "Text field_1" at 380,23 size 38x22; Text 'N/A'
   TextField "Text field_2" at 506,23 size 38x22; Text 'N/A'
   Group "Group" at 338,20 size 754x28
   Button "Open Popup" at 2,20 size 1090x28; TextOff 'Text'
   Group "Group_1" at 2,20 size 1090x28
   Rectangle "Rectangle_7" at 338,20 size 754x28
      Visibility <- "Data_Connection.DisableRecipeControl"
   TextField "Text field_3" at 629,23 size 223x23; Text 'Recipe Control Disabled / Rezepturverwaltung deaktiviert'
      Visibility <- "Data_Connection.DisableRecipeControl"
   Rectangle "Rectangle_8" at 2,20 size 1090x28
      Visibility <- "DISABLED"
   TextField "Text field_4" at 475,23 size 188x23; Text 'No Recipe Available / Kein Datensatz vorhanden'
      Visibility <- "DISABLED"
*)